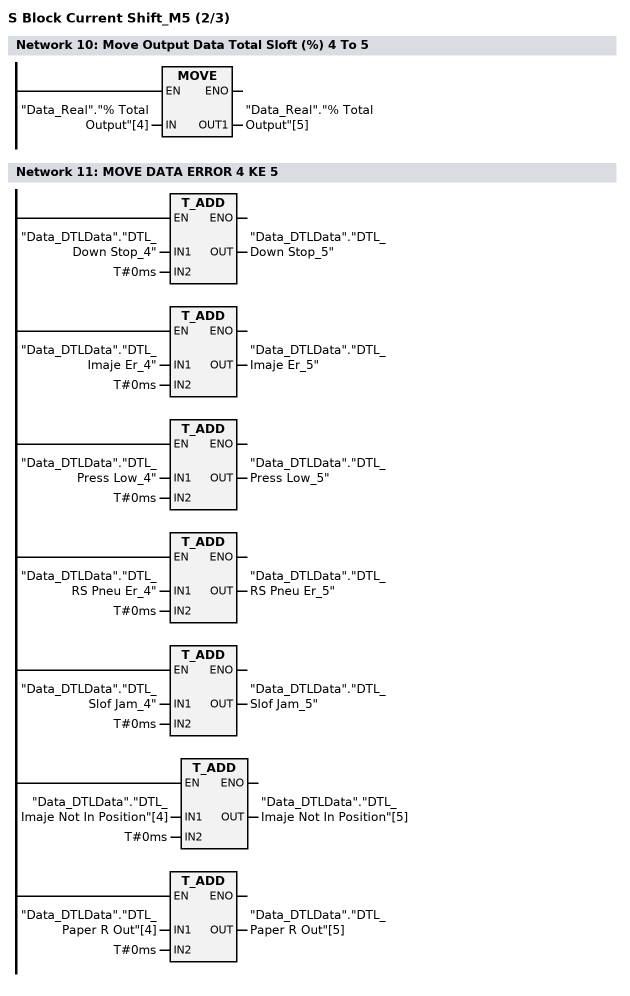
   RUNG wire#powerrail
      { S7_GenerateENO := "TRUE" } Move(in := "Data_Real"."% Total Output"[4], out1 => "Data_Real"."% Total Output"[5])
   END_RUNG
   // the same network as SCL:
   "Data_Real"."% Total Output"[5] := "Data_Real"."% Total Output"[4];
END_REGION

REGION Network 11: MOVE DATA ERROR 4 KE 5
   "Data_DTLData"."DTL_Down Stop_5" := T_ADD(IN1 := "Data_DTLData"."DTL_Down Stop_4", IN2 := T#0ms);
   "Data_DTLData"."DTL_Imaje Er_5" := T_ADD(IN1 := "Data_DTLData"."DTL_Imaje Er_4", IN2 := T#0ms);
   "Data_DTLData"."DTL_Press Low_5" := T_ADD(IN1 := "Data_DTLData"."DTL_Press Low_4", IN2 := T#0ms);
   "Data_DTLData"."DTL_RS Pneu Er_5" := T_ADD(IN1 := "Data_DTLData"."DTL_RS Pneu Er_4", IN2 := T#0ms);
   "Data_DTLData"."DTL_Slof Jam_5" := T_ADD(IN1 := "Data_DTLData"."DTL_Slof Jam_4", IN2 := T#0ms);
   "Data_DTLData"."DTL_Imaje Not In Position"[5] := T_ADD(IN1 := "Data_DTLData"."DTL_Imaje Not In Position"[4],
                           IN2 := T#0ms);
   "Data_DTLData"."DTL_Paper R Out"[5] := T_ADD(IN1 := "Data_DTLData"."DTL_Paper R Out"[4], IN2 := T#0ms);
END_REGION

REGION Network 12: Copi data frekuensi error
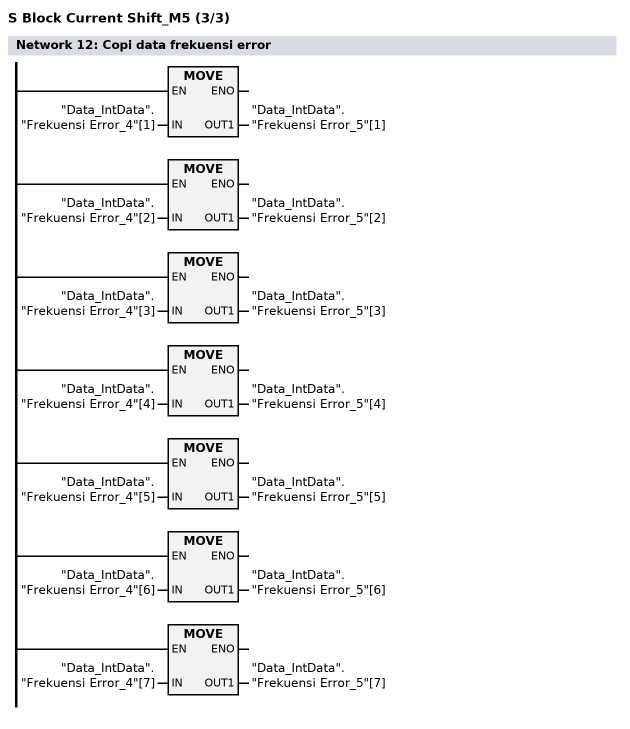
   RUNG wire#powerrail
      { S7_GenerateENO := "TRUE" } Move(in := "Data_IntData"."Frekuensi Error_4"[1], out1 => "Data_IntData"."Frekuensi Error_5"[1])
   END_RUNG
   RUNG wire#powerrail
      { S7_GenerateENO := "TRUE" } Move(in := "Data_IntData"."Frekuensi Error_4"[2], out1 => "Data_IntData"."Frekuensi Error_5"[2])
   END_RUNG
   RUNG wire#powerrail
      { S7_GenerateENO := "TRUE" } Move(in := "Data_IntData"."Frekuensi Error_4"[3], out1 => "Data_IntData"."Frekuensi Error_5"[3])
   END_RUNG
   RUNG wire#powerrail
      { S7_GenerateENO := "TRUE" } Move(in := "Data_IntData"."Frekuensi Error_4"[4], out1 => "Data_IntData"."Frekuensi Error_5"[4])
   END_RUNG
   RUNG wire#powerrail
      { S7_GenerateENO := "TRUE" } Move(in := "Data_IntData"."Frekuensi Error_4"[5], out1 => "Data_IntData"."Frekuensi Error_5"[5])
   END_RUNG
   RUNG wire#powerrail
      { S7_GenerateENO := "TRUE" } Move(in := "Data_IntData"."Frekuensi Error_4"[6], out1 => "Data_IntData"."Frekuensi Error_5"[6])
   END_RUNG
   RUNG wire#powerrail
      { S7_GenerateENO := "TRUE" } Move(in := "Data_IntData"."Frekuensi Error_4"[7], out1 => "Data_IntData"."Frekuensi Error_5"[7])
   END_RUNG
   // the same network as SCL:
   "Data_IntData"."Frekuensi Error_5"[1] := "Data_IntData"."Frekuensi Error_4"[1];
   "Data_IntData"."Frekuensi Error_5"[2] := "Data_IntData"."Frekuensi Error_4"[2];
   "Data_IntData"."Frekuensi Error_5"[3] := "Data_IntData"."Frekuensi Error_4"[3];
   "Data_IntData"."Frekuensi Error_5"[4] := "Data_IntData"."Frekuensi Error_4"[4];
   "Data_IntData"."Frekuensi Error_5"[5] := "Data_IntData"."Frekuensi Error_4"[5];
   "Data_IntData"."Frekuensi Error_5"[6] := "Data_IntData"."Frekuensi Error_4"[6];
   "Data_IntData"."Frekuensi Error_5"[7] := "Data_IntData"."Frekuensi Error_4"[7];
END_REGION
END_FUNCTION_BLOCK

FUNCTION "RS 1 Pneumatic Pusher Advance" : Void   // FC1, LAD
{ S7_Optimized_Access := 'TRUE' }
VERSION : 0.1
BEGIN

REGION Network 1: Reed Switch Pneumatic 1 Advance Error
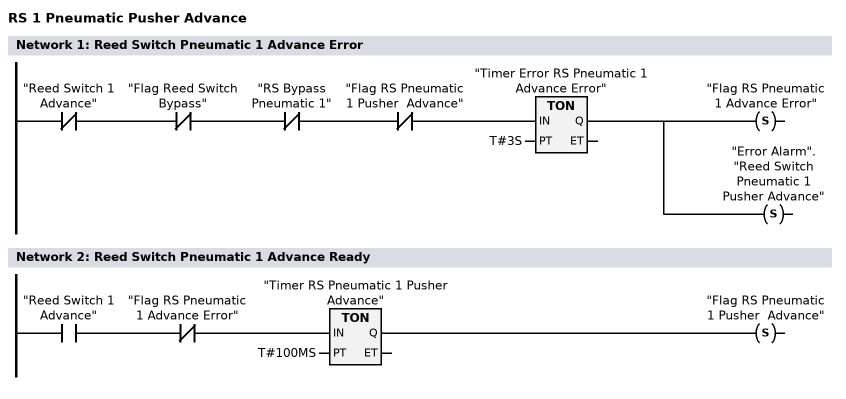
   "Timer Error RS Pneumatic 1 Advance Error".TON(IN := NOT "Reed Switch 1 Advance" AND NOT "Flag Reed Switch Bypass" AND NOT "RS Bypass Pneumatic 1" AND NOT "Flag RS Pneumatic 1 Pusher  Advance",
                           PT := T#3S);
   IF "Timer Error RS Pneumatic 1 Advance Error".Q THEN
       "Flag RS Pneumatic 1 Advance Error" := TRUE;
       "Error Alarm"."Reed Switch Pneumatic 1 Pusher Advance" := TRUE;
   END_IF;
END_REGION

REGION Network 2: Reed Switch Pneumatic 1 Advance Ready
   "Timer RS Pneumatic 1 Pusher Advance".TON(IN := "Reed Switch 1 Advance" AND NOT "Flag RS Pneumatic 1 Advance Error",
                           PT := T#100MS);
   IF "Timer RS Pneumatic 1 Pusher Advance".Q THEN "Flag RS Pneumatic 1 Pusher  Advance" := TRUE; END_IF;
END_REGION
END_FUNCTION

FUNCTION "RS 2 Pneumatic Pusher Retract" : Void   // FC2, LAD
{ S7_Optimized_Access := 'TRUE' }
VERSION : 0.1
BEGIN

REGION Network 1: Reed Switch Pneumatic 1 Upper Error
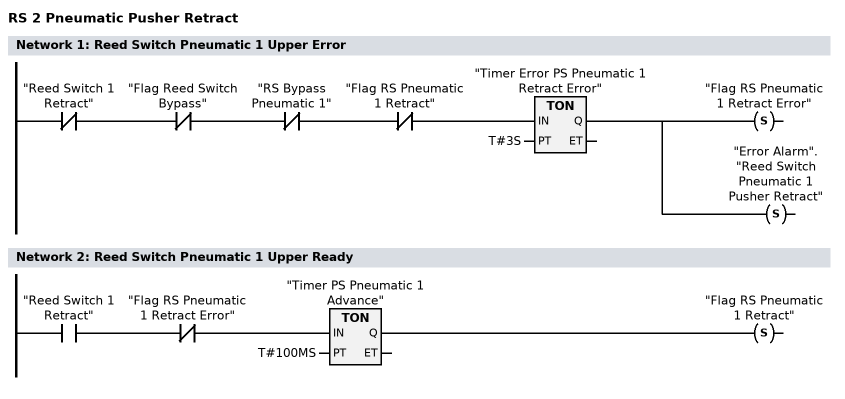
   "Timer Error PS Pneumatic 1 Retract Error".TON(IN := NOT "Reed Switch 1 Retract" AND NOT "Flag Reed Switch Bypass" AND NOT "RS Bypass Pneumatic 1" AND NOT "Flag RS Pneumatic 1 Retract",
                           PT := T#3S);
   IF "Timer Error PS Pneumatic 1 Retract Error".Q THEN
       "Flag RS Pneumatic 1 Retract Error" := TRUE;
       "Error Alarm"."Reed Switch Pneumatic 1 Pusher Retract" := TRUE;
   END_IF;
END_REGION

REGION Network 2: Reed Switch Pneumatic 1 Upper Ready
   "Timer PS Pneumatic 1 Advance".TON(IN := "Reed Switch 1 Retract" AND NOT "Flag RS Pneumatic 1 Retract Error",
                           PT := T#100MS);
   IF "Timer PS Pneumatic 1 Advance".Q THEN "Flag RS Pneumatic 1 Retract" := TRUE; END_IF;
END_REGION
END_FUNCTION

FUNCTION "RS 3 Pneumatic 3 Up" : Void   // FC3, LAD
{ S7_Optimized_Access := 'TRUE' }
VERSION : 0.1
BEGIN

REGION Network 1: Reed Switch Pneumatic 3 Up Error
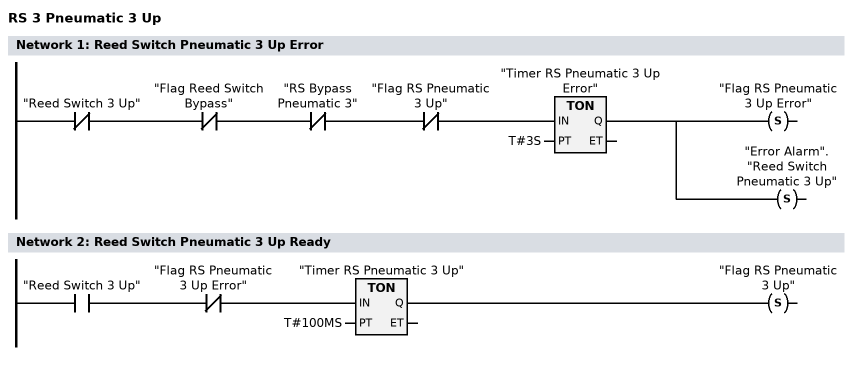
   "Timer RS Pneumatic 3 Up Error".TON(IN := NOT "Reed Switch 3 Up" AND NOT "Flag Reed Switch Bypass" AND NOT "RS Bypass Pneumatic 3" AND NOT "Flag RS Pneumatic 3 Up",
                           PT := T#3S);
   IF "Timer RS Pneumatic 3 Up Error".Q THEN
       "Flag RS Pneumatic 3 Up Error" := TRUE;
       "Error Alarm"."Reed Switch Pneumatic 3 Up" := TRUE;
   END_IF;
END_REGION

REGION Network 2: Reed Switch Pneumatic 3 Up Ready
   "Timer RS Pneumatic 3 Up".TON(IN := "Reed Switch 3 Up" AND NOT "Flag RS Pneumatic 3 Up Error", PT := T#100MS);
   IF "Timer RS Pneumatic 3 Up".Q THEN "Flag RS Pneumatic 3 Up" := TRUE; END_IF;
END_REGION
END_FUNCTION

FUNCTION "RS 4 Pneumatic 3 Down" : Void   // FC4, LAD
{ S7_Optimized_Access := 'TRUE' }
VERSION : 0.1
BEGIN

REGION Network 1: Reed Switch Pneumatic 3 Down Error
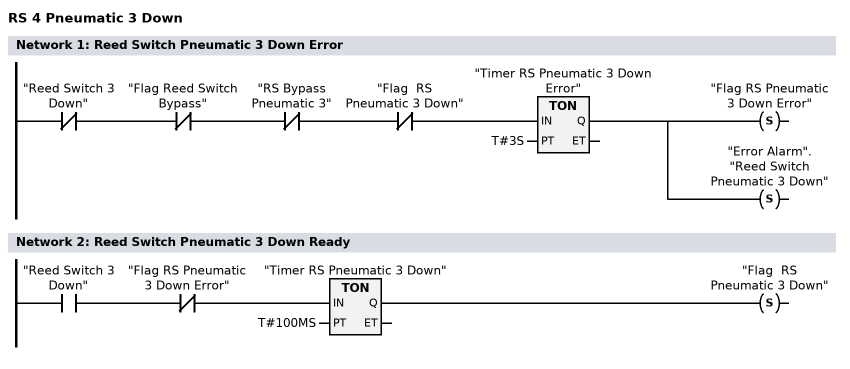
   "Timer RS Pneumatic 3 Down Error".TON(IN := NOT "Reed Switch 3 Down" AND NOT "Flag Reed Switch Bypass" AND NOT "RS Bypass Pneumatic 3" AND NOT "Flag  RS Pneumatic 3 Down",
                           PT := T#3S);
   IF "Timer RS Pneumatic 3 Down Error".Q THEN
       "Flag RS Pneumatic 3 Down Error" := TRUE;
       "Error Alarm"."Reed Switch Pneumatic 3 Down" := TRUE;
   END_IF;
END_REGION

REGION Network 2: Reed Switch Pneumatic 3 Down Ready
   "Timer RS Pneumatic 3 Down".TON(IN := "Reed Switch 3 Down" AND NOT "Flag RS Pneumatic 3 Down Error",
                           PT := T#100MS);
   IF "Timer RS Pneumatic 3 Down".Q THEN "Flag  RS Pneumatic 3 Down" := TRUE; END_IF;
END_REGION
END_FUNCTION

FUNCTION "RS 5 Pneumatic 4 Down" : Void   // FC5, LAD
{ S7_Optimized_Access := 'TRUE' }
VERSION : 0.1
BEGIN

REGION Network 1: Reed Switch Pneumatic 4 Down Error
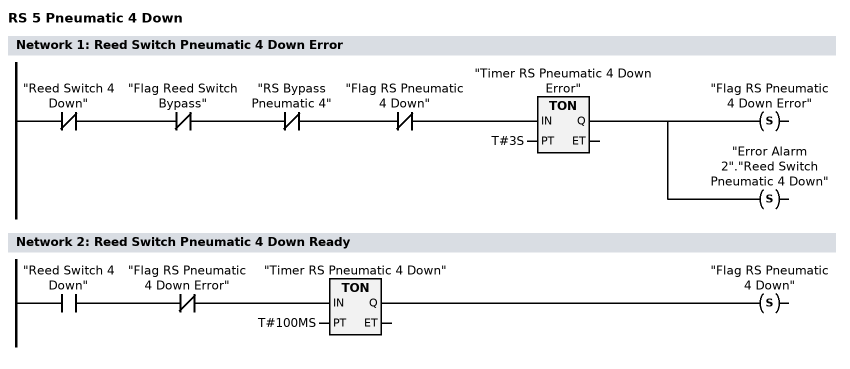
   "Timer RS Pneumatic 4 Down Error".TON(IN := NOT "Reed Switch 4 Down" AND NOT "Flag Reed Switch Bypass" AND NOT "RS Bypass Pneumatic 4" AND NOT "Flag RS Pneumatic 4 Down",
                           PT := T#3S);
   IF "Timer RS Pneumatic 4 Down Error".Q THEN
       "Flag RS Pneumatic 4 Down Error" := TRUE;
       "Error Alarm 2"."Reed Switch Pneumatic 4 Down" := TRUE;
   END_IF;
END_REGION

REGION Network 2: Reed Switch Pneumatic 4 Down Ready
   "Timer RS Pneumatic 4 Down".TON(IN := "Reed Switch 4 Down" AND NOT "Flag RS Pneumatic 4 Down Error",
                           PT := T#100MS);
   IF "Timer RS Pneumatic 4 Down".Q THEN "Flag RS Pneumatic 4 Down" := TRUE; END_IF;
END_REGION
END_FUNCTION

FUNCTION "RS 6 Pneumatic 4 Up" : Void   // FC6, LAD
{ S7_Optimized_Access := 'TRUE' }
VERSION : 0.1
BEGIN

REGION Network 1: Reed Switch Pneumatic 4 Up Error
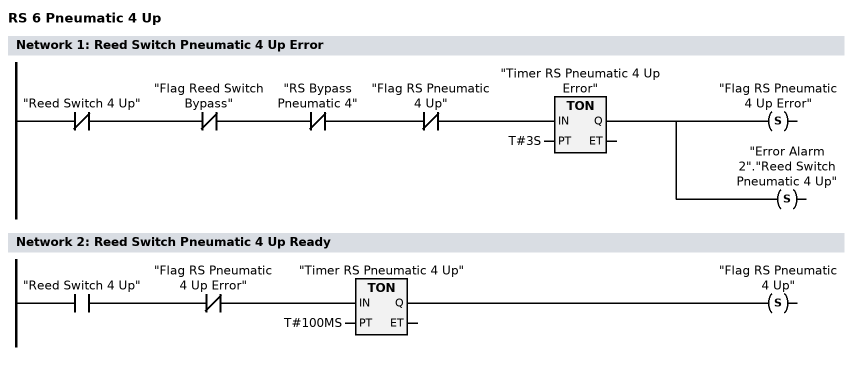
   "Timer RS Pneumatic 4 Up Error".TON(IN := NOT "Reed Switch 4 Up" AND NOT "Flag Reed Switch Bypass" AND NOT "RS Bypass Pneumatic 4" AND NOT "Flag RS Pneumatic 4 Up",
                           PT := T#3S);
   IF "Timer RS Pneumatic 4 Up Error".Q THEN
       "Flag RS Pneumatic 4 Up Error" := TRUE;
       "Error Alarm 2"."Reed Switch Pneumatic 4 Up" := TRUE;
   END_IF;
END_REGION

REGION Network 2: Reed Switch Pneumatic 4 Up Ready
   "Timer RS Pneumatic 4 Up".TON(IN := "Reed Switch 4 Up" AND NOT "Flag RS Pneumatic 4 Up Error", PT := T#100MS);
   IF "Timer RS Pneumatic 4 Up".Q THEN "Flag RS Pneumatic 4 Up" := TRUE; END_IF;
END_REGION
END_FUNCTION

FUNCTION "RS 7 Pneumatic 5 Advance" : Void   // FC7, LAD
{ S7_Optimized_Access := 'TRUE' }
VERSION : 0.1
BEGIN

REGION Network 1: Reed Switch Pneumatic 5 Advance Error
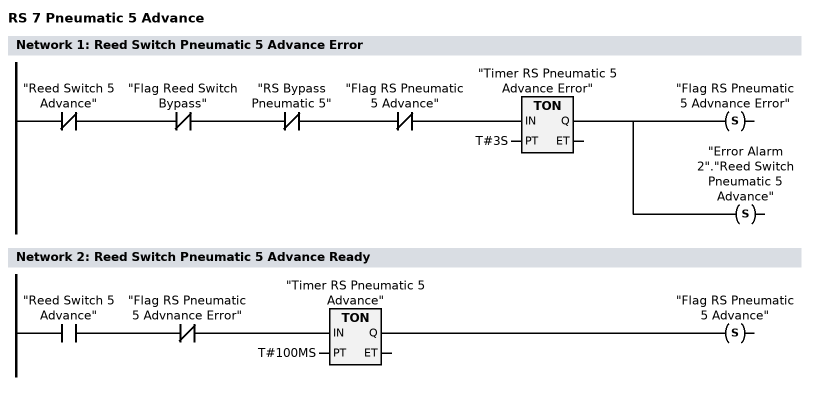
   "Timer RS Pneumatic 5 Advance Error".TON(IN := NOT "Reed Switch 5 Advance" AND NOT "Flag Reed Switch Bypass" AND NOT "RS Bypass Pneumatic 5" AND NOT "Flag RS Pneumatic 5 Advance",
                           PT := T#3S);
   IF "Timer RS Pneumatic 5 Advance Error".Q THEN
       "Flag RS Pneumatic 5 Advnance Error" := TRUE;
       "Error Alarm 2"."Reed Switch Pneumatic 5 Advance" := TRUE;
   END_IF;
END_REGION

REGION Network 2: Reed Switch Pneumatic 5 Advance Ready
   "Timer RS Pneumatic 5 Advance".TON(IN := "Reed Switch 5 Advance" AND NOT "Flag RS Pneumatic 5 Advnance Error",
                           PT := T#100MS);
   IF "Timer RS Pneumatic 5 Advance".Q THEN "Flag RS Pneumatic 5 Advance" := TRUE; END_IF;
END_REGION
END_FUNCTION

FUNCTION "RS 8 Pneumatic 5 Retract" : Void   // FC8, LAD
{ S7_Optimized_Access := 'TRUE' }
VERSION : 0.1
BEGIN

REGION Network 1: Reed Switch Pneumatic 5 Retract Error
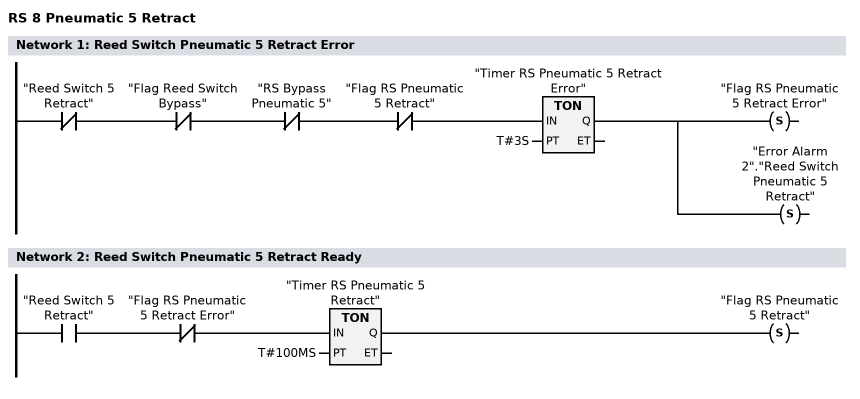
   "Timer RS Pneumatic 5 Retract Error".TON(IN := NOT "Reed Switch 5 Retract" AND NOT "Flag Reed Switch Bypass" AND NOT "RS Bypass Pneumatic 5" AND NOT "Flag RS Pneumatic 5 Retract",
                           PT := T#3S);
   IF "Timer RS Pneumatic 5 Retract Error".Q THEN
       "Flag RS Pneumatic 5 Retract Error" := TRUE;
       "Error Alarm 2"."Reed Switch Pneumatic 5 Retract" := TRUE;
   END_IF;
END_REGION

REGION Network 2: Reed Switch Pneumatic 5 Retract Ready
   "Timer RS Pneumatic 5 Retract".TON(IN := "Reed Switch 5 Retract" AND NOT "Flag RS Pneumatic 5 Retract Error",
                           PT := T#100MS);
   IF "Timer RS Pneumatic 5 Retract".Q THEN "Flag RS Pneumatic 5 Retract" := TRUE; END_IF;
END_REGION
END_FUNCTION

ORGANIZATION_BLOCK "Main"   // OB1, LAD, ProgramCycle
TITLE = "Main Program Sweep (Cycle)"
{ S7_Optimized_Access := 'TRUE' }
VERSION : 0.1
   VAR_TEMP   // added for the SCL form of the ladder/FBD networks
      _w1 : Bool;
      _w2 : Bool;
      _w3 : Bool;
      _w4 : Bool;
      _w5 : Bool;
   END_VAR
BEGIN

REGION Network 1: Machine Stand by
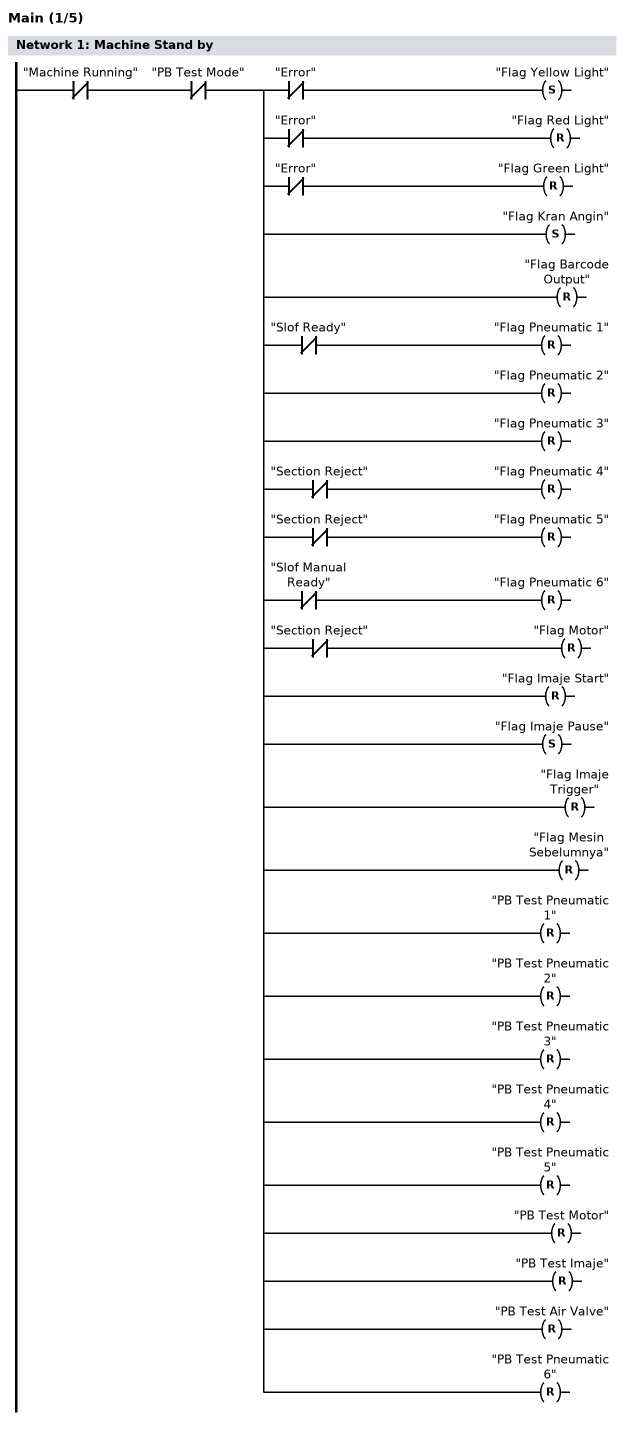
   RUNG wire#powerrail
      I_Contact( "Machine Running" )
      I_Contact( "PB Test Mode" )
      wire#w1
      I_Contact( "Error" )
      S_Coil( "Flag Yellow Light" )
   END_RUNG
   RUNG wire#w1
      I_Contact( "Error" )
      R_Coil( "Flag Red Light" )
   END_RUNG
   RUNG wire#w1
      I_Contact( "Error" )
      R_Coil( "Flag Green Light" )
   END_RUNG
   RUNG wire#w1
      S_Coil( "Flag Kran Angin" )
   END_RUNG
   RUNG wire#w1
      R_Coil( "Flag Barcode Output" )
   END_RUNG
   RUNG wire#w1
      I_Contact( "Slof Ready" )
      R_Coil( "Flag Pneumatic 1" )
   END_RUNG
   RUNG wire#w1
      R_Coil( "Flag Pneumatic 2" )
   END_RUNG
   RUNG wire#w1
      R_Coil( "Flag Pneumatic 3" )
   END_RUNG
   RUNG wire#w1
      I_Contact( "Section Reject" )
      R_Coil( "Flag Pneumatic 4" )
   END_RUNG
   RUNG wire#w1
      I_Contact( "Section Reject" )
      R_Coil( "Flag Pneumatic 5" )
   END_RUNG
   RUNG wire#w1
      I_Contact( "Slof Manual Ready" )
      R_Coil( "Flag Pneumatic 6" )
   END_RUNG
   RUNG wire#w1
      I_Contact( "Section Reject" )
      R_Coil( "Flag Motor" )
   END_RUNG
   RUNG wire#w1
      R_Coil( "Flag Imaje Start" )
   END_RUNG
   RUNG wire#w1
      S_Coil( "Flag Imaje Pause" )
   END_RUNG
   RUNG wire#w1
      R_Coil( "Flag Imaje Trigger" )
   END_RUNG
   RUNG wire#w1
      R_Coil( "Flag Mesin Sebelumnya" )
   END_RUNG
   RUNG wire#w1
      R_Coil( "PB Test Pneumatic 1" )
   END_RUNG
   RUNG wire#w1
      R_Coil( "PB Test Pneumatic 2" )
   END_RUNG
   RUNG wire#w1
      R_Coil( "PB Test Pneumatic 3" )
   END_RUNG
   RUNG wire#w1
      R_Coil( "PB Test Pneumatic 4" )
   END_RUNG
   RUNG wire#w1
      R_Coil( "PB Test Pneumatic 5" )
   END_RUNG
   RUNG wire#w1
      R_Coil( "PB Test Motor" )
   END_RUNG
   RUNG wire#w1
      R_Coil( "PB Test Imaje" )
   END_RUNG
   RUNG wire#w1
      R_Coil( "PB Test Air Valve" )
   END_RUNG
   RUNG wire#w1
      R_Coil( "PB Test Pneumatic 6" )
   END_RUNG
   // the same network as SCL:
   #_w1 := NOT "Machine Running" AND NOT "PB Test Mode";
   IF #_w1 AND NOT "Error" THEN
       "Flag Yellow Light" := TRUE;
       "Flag Red Light" := FALSE;
       "Flag Green Light" := FALSE;
   END_IF;
   IF #_w1 THEN
       "Flag Kran Angin" := TRUE;
       "Flag Barcode Output" := FALSE;
   END_IF;
   IF #_w1 AND NOT "Slof Ready" THEN "Flag Pneumatic 1" := FALSE; END_IF;
   IF #_w1 THEN
       "Flag Pneumatic 2" := FALSE;
       "Flag Pneumatic 3" := FALSE;
   END_IF;
   IF #_w1 AND NOT "Section Reject" THEN
       "Flag Pneumatic 4" := FALSE;
       "Flag Pneumatic 5" := FALSE;
   END_IF;
   IF #_w1 AND NOT "Slof Manual Ready" THEN "Flag Pneumatic 6" := FALSE; END_IF;
   IF #_w1 AND NOT "Section Reject" THEN "Flag Motor" := FALSE; END_IF;
   IF #_w1 THEN
       "Flag Imaje Start" := FALSE;
       "Flag Imaje Pause" := TRUE;
       "Flag Imaje Trigger" := FALSE;
       "Flag Mesin Sebelumnya" := FALSE;
       "PB Test Pneumatic 1" := FALSE;
       "PB Test Pneumatic 2" := FALSE;
       "PB Test Pneumatic 3" := FALSE;
       "PB Test Pneumatic 4" := FALSE;
       "PB Test Pneumatic 5" := FALSE;
       "PB Test Motor" := FALSE;
       "PB Test Imaje" := FALSE;
       "PB Test Air Valve" := FALSE;
       "PB Test Pneumatic 6" := FALSE;
   END_IF;
END_REGION

REGION Network 2: Output
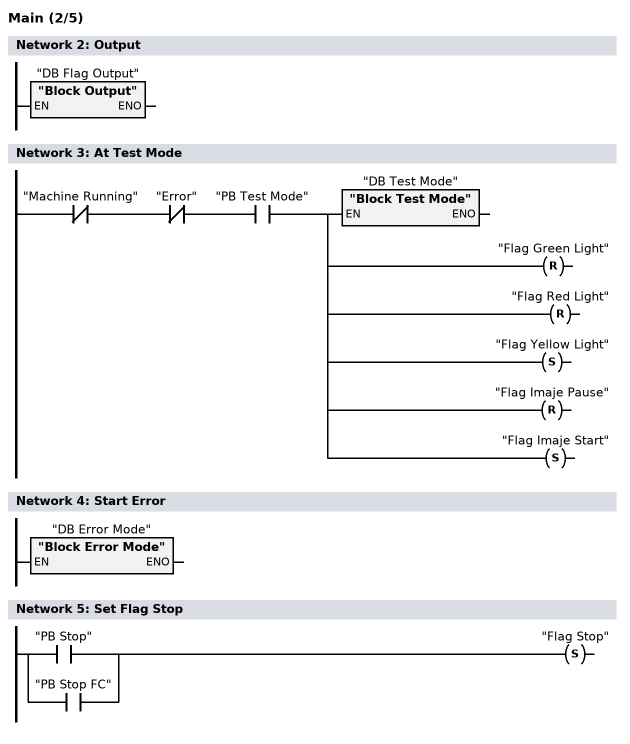
   RUNG wire#powerrail
      "DB Flag Output"()
   END_RUNG
   // the same network as SCL:
   "DB Flag Output"();   // "Block Output"
END_REGION

REGION Network 3: At Test Mode
   RUNG wire#powerrail
      I_Contact( "Machine Running" )
      I_Contact( "Error" )
      Contact( "PB Test Mode" )
      wire#w1
      "DB Test Mode"()
   END_RUNG
   RUNG wire#w1
      R_Coil( "Flag Green Light" )
   END_RUNG
   RUNG wire#w1
      R_Coil( "Flag Red Light" )
   END_RUNG
   RUNG wire#w1
      S_Coil( "Flag Yellow Light" )
   END_RUNG
   RUNG wire#w1
      R_Coil( "Flag Imaje Pause" )
   END_RUNG
   RUNG wire#w1
      S_Coil( "Flag Imaje Start" )
   END_RUNG
   // the same network as SCL:
   #_w1 := NOT "Machine Running" AND NOT "Error" AND "PB Test Mode";
   IF #_w1 THEN
       "DB Test Mode"();   // "Block Test Mode"
       "Flag Green Light" := FALSE;
       "Flag Red Light" := FALSE;
       "Flag Yellow Light" := TRUE;
       "Flag Imaje Pause" := FALSE;
       "Flag Imaje Start" := TRUE;
   END_IF;
END_REGION

REGION Network 4: Start Error
   RUNG wire#powerrail
      "DB Error Mode"()
   END_RUNG
   // the same network as SCL:
   "DB Error Mode"();   // "Block Error Mode"
END_REGION

REGION Network 5: Set Flag Stop
   RUNG wire#powerrail
      Contact( "PB Stop" )
      wire#w1
      S_Coil( "Flag Stop" )
   END_RUNG
   RUNG wire#powerrail
      Contact( "PB Stop FC" )
   END_RUNG wire#w1
   // the same network as SCL:
   IF "PB Stop" OR "PB Stop FC" THEN "Flag Stop" := TRUE; END_IF;
END_REGION

REGION Network 6: Flag Stop
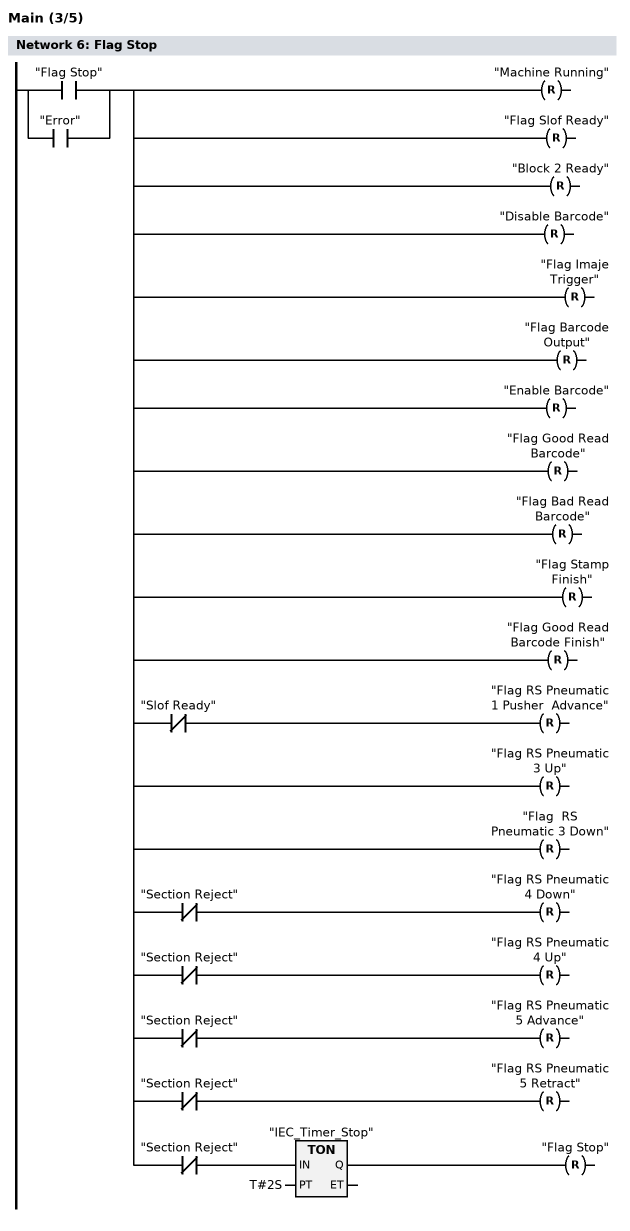
   #_w1 := "Flag Stop" OR "Error";
   IF #_w1 THEN
       "Machine Running" := FALSE;
       "Flag Slof Ready" := FALSE;
       "Block 2 Ready" := FALSE;
       "Disable Barcode" := FALSE;
       "Flag Imaje Trigger" := FALSE;
       "Flag Barcode Output" := FALSE;
       "Enable Barcode" := FALSE;
       "Flag Good Read Barcode" := FALSE;
       "Flag Bad Read Barcode" := FALSE;
       "Flag Stamp Finish" := FALSE;
       "Flag Good Read Barcode Finish" := FALSE;
   END_IF;
   IF #_w1 AND NOT "Slof Ready" THEN "Flag RS Pneumatic 1 Pusher  Advance" := FALSE; END_IF;
   IF #_w1 THEN
       "Flag RS Pneumatic 3 Up" := FALSE;
       "Flag  RS Pneumatic 3 Down" := FALSE;
   END_IF;
   IF #_w1 AND NOT "Section Reject" THEN
       "Flag RS Pneumatic 4 Down" := FALSE;
       "Flag RS Pneumatic 4 Up" := FALSE;
       "Flag RS Pneumatic 5 Advance" := FALSE;
       "Flag RS Pneumatic 5 Retract" := FALSE;
   END_IF;
   "IEC_Timer_Stop".TON(IN := #_w1 AND NOT "Section Reject", PT := T#2S);
   IF "IEC_Timer_Stop".Q THEN "Flag Stop" := FALSE; END_IF;
END_REGION

REGION Network 7: PB Run
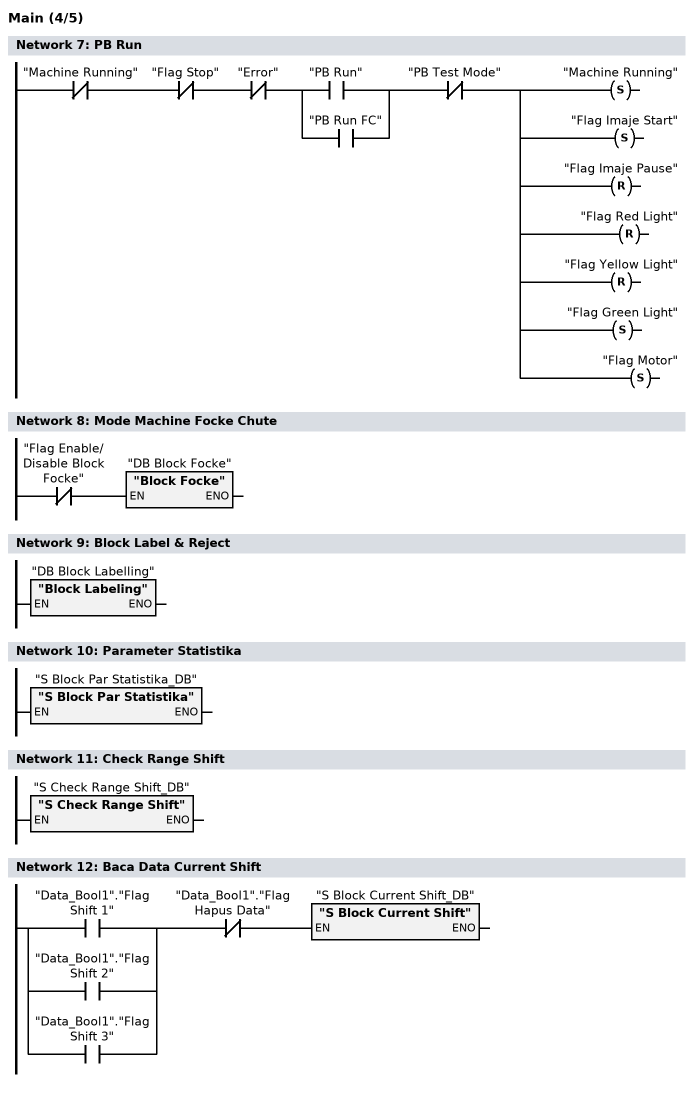
   RUNG wire#powerrail
      I_Contact( "Machine Running" )
      I_Contact( "Flag Stop" )
      I_Contact( "Error" )
      wire#w1
      Contact( "PB Run" )
      wire#w2
      I_Contact( "PB Test Mode" )
      wire#w3
      S_Coil( "Machine Running" )
   END_RUNG
   RUNG wire#w1
      Contact( "PB Run FC" )
   END_RUNG wire#w2
   RUNG wire#w3
      S_Coil( "Flag Imaje Start" )
   END_RUNG
   RUNG wire#w3
      R_Coil( "Flag Imaje Pause" )
   END_RUNG
   RUNG wire#w3
      R_Coil( "Flag Red Light" )
   END_RUNG
   RUNG wire#w3
      R_Coil( "Flag Yellow Light" )
   END_RUNG
   RUNG wire#w3
      S_Coil( "Flag Green Light" )
   END_RUNG
   RUNG wire#w3
      S_Coil( "Flag Motor" )
   END_RUNG
   // the same network as SCL:
   #_w1 := NOT "Machine Running" AND NOT "Flag Stop" AND NOT "Error" AND ("PB Run" OR "PB Run FC") AND NOT "PB Test Mode";
   IF #_w1 THEN
       "Machine Running" := TRUE;
       "Flag Imaje Start" := TRUE;
       "Flag Imaje Pause" := FALSE;
       "Flag Red Light" := FALSE;
       "Flag Yellow Light" := FALSE;
       "Flag Green Light" := TRUE;
       "Flag Motor" := TRUE;
   END_IF;
END_REGION

REGION Network 8: Mode Machine Focke Chute
   RUNG wire#powerrail
      I_Contact( "Flag Enable/Disable Block Focke" )
      "DB Block Focke"()
   END_RUNG
   // the same network as SCL:
   IF NOT "Flag Enable/Disable Block Focke" THEN
       "DB Block Focke"();   // "Block Focke"
   END_IF;
END_REGION

REGION Network 9: Block Label & Reject
   RUNG wire#powerrail
      "DB Block Labelling"()
   END_RUNG
   // the same network as SCL:
   "DB Block Labelling"();   // "Block Labeling"
END_REGION

REGION Network 10: Parameter Statistika
   RUNG wire#powerrail
      "S Block Par Statistika_DB"()
   END_RUNG
   // the same network as SCL:
   "S Block Par Statistika_DB"();   // "S Block Par Statistika"
END_REGION

REGION Network 11: Check Range Shift
   RUNG wire#powerrail
      "S Check Range Shift_DB"()
   END_RUNG
   // the same network as SCL:
   "S Check Range Shift_DB"();   // "S Check Range Shift"
END_REGION

REGION Network 12: Baca Data Current Shift
   RUNG wire#powerrail
      Contact( "Data_Bool1"."Flag Shift 1" )
      wire#w1
      I_Contact( "Data_Bool1"."Flag Hapus Data" )
      "S Block Current Shift_DB"()
   END_RUNG
   RUNG wire#powerrail
      Contact( "Data_Bool1"."Flag Shift 2" )
   END_RUNG wire#w1
   RUNG wire#powerrail
      Contact( "Data_Bool1"."Flag Shift 3" )
   END_RUNG wire#w1
   // the same network as SCL:
   IF ("Data_Bool1"."Flag Shift 1" OR "Data_Bool1"."Flag Shift 2" OR "Data_Bool1"."Flag Shift 3") AND NOT "Data_Bool1"."Flag Hapus Data" THEN
       "S Block Current Shift_DB"();   // "S Block Current Shift"
   END_IF;
END_REGION

REGION Network 13: Copi Data Jika Power Mati Pada Waktu Proses Pindah Data (Belum ada)
END_REGION

REGION Network 14: Copy Data Current Shift Min 1 Sampai Min 5 Dan Hapus Data